      Carrier64_Faults_1 : Int := 238;
      Carrier64_Faults_2 : Int := 239;
      Carrier64_Faults_3 : Int := 240;
      Carrier65_Faults_0 : Int := 241;
      Carrier65_Faults_1 : Int := 242;
      Carrier65_Faults_2 : Int := 243;
      Carrier65_Faults_3 : Int := 244;
      Carrier66_Faults_0 : Int := 245;
      Carrier66_Faults_1 : Int := 246;
      Carrier66_Faults_2 : Int := 247;
      Carrier66_Faults_3 : Int := 248;
      Carrier67_Faults_0 : Int := 249;
      Carrier67_Faults_1 : Int := 250;
      Carrier67_Faults_2 : Int := 251;
      Carrier67_Faults_3 : Int := 252;
      Carrier68_Faults_0 : Int := 253;
      Carrier68_Faults_1 : Int := 254;
      Carrier68_Faults_2 : Int := 255;
      Carrier68_Faults_3 : Int := 256;
      Carrier69_Faults_0 : Int := 257;
      Carrier69_Faults_1 : Int := 258;
      Carrier69_Faults_2 : Int := 259;
      Carrier69_Faults_3 : Int := 260;
      Carrier70_Faults_0 : Int := 261;
      Carrier70_Faults_1 : Int := 262;
      Carrier70_Faults_2 : Int := 263;
      Carrier70_Faults_3 : Int := 264;
      Carrier71_Faults_0 : Int := 265;
      Carrier71_Faults_1 : Int := 266;
      Carrier71_Faults_2 : Int := 267;
      Carrier71_Faults_3 : Int := 268;
      Carrier72_Faults_0 : Int := 269;
      Carrier72_Faults_1 : Int := 270;
      Carrier72_Faults_2 : Int := 271;
      Carrier72_Faults_3 : Int := 272;
      Carrier73_Faults_0 : Int := 273;
      Carrier73_Faults_1 : Int := 274;
      Carrier73_Faults_2 : Int := 275;
      Carrier73_Faults_3 : Int := 276;
      Carrier74_Faults_0 : Int := 277;
      Carrier74_Faults_1 : Int := 278;
      Carrier74_Faults_2 : Int := 279;
      Carrier74_Faults_3 : Int := 280;
      Carrier75_Faults_0 : Int := 281;
      Carrier75_Faults_1 : Int := 282;
      Carrier75_Faults_2 : Int := 283;
      Carrier75_Faults_3 : Int := 284;
      Carrier76_Faults_0 : Int := 285;
      Carrier76_Faults_1 : Int := 286;
      Carrier76_Faults_2 : Int := 287;
      Carrier76_Faults_3 : Int := 288;
      Carrier77_Faults_0 : Int := 289;
      Carrier77_Faults_1 : Int := 290;
      Carrier77_Faults_2 : Int := 291;
      Carrier77_Faults_3 : Int := 292;
      Carrier78_Faults_0 : Int := 293;
      Carrier78_Faults_1 : Int := 294;
      Carrier78_Faults_2 : Int := 295;
      Carrier78_Faults_3 : Int := 296;
      Carrier79_Faults_0 : Int := 297;
      Carrier79_Faults_1 : Int := 298;
      Carrier79_Faults_2 : Int := 299;
      Carrier79_Faults_3 : Int := 300;
      Carrier80_Faults_0 : Int := 301;
      Carrier80_Faults_1 : Int := 302;
      Carrier80_Faults_2 : Int := 303;
      Carrier80_Faults_3 : Int := 304;
      Carrier81_Faults_0 : Int := 305;
      Carrier81_Faults_1 : Int := 306;
      Carrier81_Faults_2 : Int := 307;
      Carrier81_Faults_3 : Int := 308;
      Carrier82_Faults_0 : Int := 309;
      Carrier82_Faults_1 : Int := 310;
      Carrier82_Faults_2 : Int := 311;
      Carrier82_Faults_3 : Int := 312;
   END_VAR
BEGIN
END_DATA_BLOCK

DATA_BLOCK "DB401_HMI_Status"   // DB401
{ S7_Optimized_Access := 'TRUE' }
VERSION : 0.1
   VAR
      Drive : "UDT_Drive_HMI";
      IO : "UDT_Carrier_IO_HMI";
      Status : "UDT_Carrier_Status_HMI";
      ZoneStatus : "UDT_Zone_Status_HMI";
   END_VAR
BEGIN
END_DATA_BLOCK

DATA_BLOCK "DB402_SDC_CARRIER_DRIVE_DATA"   // DB402
{ S7_Optimized_Access := 'TRUE' }
VERSION : 0.1
   VAR
      Drive_Data : "UDT_Carrier_Drive_Data";
   END_VAR
BEGIN
END_DATA_BLOCK

DATA_BLOCK "DB403_SDC_CARRIER_IO"   // DB403
{ S7_Optimized_Access := 'TRUE' }
VERSION : 0.1
   VAR
      IO_Data : "UDT_Carrier_IO_Data";
   END_VAR
BEGIN
END_DATA_BLOCK

DATA_BLOCK "Data_block_DO_NOT_CHANGE"   // DB999
{ S7_Optimized_Access := 'TRUE' }
VERSION : 0.1
   VAR RETAIN
      Production_Spacing_Memory : Int := 1000;
      Carrier_Spacing_Memory : Int := 800;
   END_VAR
BEGIN
END_DATA_BLOCK

DATA_BLOCK "DB1000_AB_Interlocks"   // DB1000
{ S7_Optimized_Access := 'TRUE' }
VERSION : 0.1
   VAR
      Interlock : "UDT_AB_Interlocks";
   END_VAR
BEGIN
END_DATA_BLOCK

DATA_BLOCK "DB_SDC_GLOBAL"   // DB3700
{ S7_Optimized_Access := 'FALSE' }
AUTHOR : FFM
FAMILY : SDC
NAME : GLOBAL
VERSION : 1.0
   VAR
      EMS_ID_ACT : Int := 130;   // Aktuelle Anzahl der EMS-Treiber
      EMS_ID_MIN : Int := 1;   // Minimum EMS ID
      EMS_ID_MAX : Int := 184;   // Maximum EMS ID
      min_barcode_mm : DInt := 900;   // Lower limit, bar code value
      max_barcode_mm : DInt := 2076000;   // Upper limit, bar code value
      START_COURSE : DInt := 5800;   // Start Barcodevalue of Course
      END_COURSE : DInt := 312200;   // Ende Barcodewert vom Kurs
      SEK_MIN : Int := 1;   // Erste Abschnitt Nummer
      SEK_MAX : Int := 508;   // Aktuelle Anzahl der Bahnabschnitte
      TAKT_TIME : Int := 0;   // Reserve
      SEK_CYCLE_COUNTER : Int := 423;   // Section for increasing the track cycle counter
      MAN_V_1 : DInt := 6000;   // manual mode, set value: drive speed (mm/min)
      MAN_V_2 : DInt := 6000;   // manual mode, set value: drive speed (mm/min)
      min_Sequence_monitor_mm : DInt := 0;   // Lower limit of bar code value for sequence monitoring
      max_Sequence_monitor_mm : DInt := 0;   // Upper limit of bar code value for sequence monitoring
      MAX_PROFIL : Int := 10;   // maximal Profil Numbers
      CURR_EMS_ID_MAX : Int := 184;   // derzeit höchsten EMS-Nummer aktiv
      current_EMS_loop : Int := 0;   // Aktuelle Anzahl der EMS-Treiber auf Schleife
      EMS_ID_BUSY : Int := 0;   // EMS Driver wird aktiviert oder deaktiviert
      TAKT_TIME_LAST : Int := 0;   // Reserve
      Reserve_56 : Array[56..59] of Byte;
      SEK_REPAIR_1 : Int := 473;   // Section for repair, reset "send to repair 1" bit
      SEK_REPAIR_2 : Int := 0;   // Section for repair, reset "send to repair 2" bit
      SEK_DIAG_1 : Int := 0;   // Section diagnosticstation 1
      SEK_DIAG_2 : Int := 0;   // Section diagnosticstation 2
      SEK_DIAG_3 : Int := 0;   // Section diagnosticstation 2
      SEK_REP_1_START : Int := 470;
      SEK_REP_1_ENDE : Int := 472;
      SEK_REP_2_START : Int := 475;
      SEK_REP_2_ENDE : Int := 475;
      INFO_REP_1_DIAG_1 : Int := 0;   // Info for Function Rep 1 at Dignosticstation 1
      INFO_REP_2_DIAG_1 : Int := 0;   // Info for Function Rep 2 at Dignosticstation 1
      INFO_REP_1_DIAG_2 : Int := 0;   // Info for Function Rep 1 at Dignosticstation 2
      INFO_REP_2_DIAG_2 : Int := 0;   // Info for Function Rep 2 at Dignosticstation 2
      INFO_REP_1_DIAG_3 : Int := 0;   // Info for Function Rep 1 at Dignosticstation 2
      INFO_REP_2_DIAG_3 : Int := 0;   // Info for Function Rep 2 at Dignosticstation 2
      EMS_VCleaner_1 : Int := 0;   // EMS mit Vaccumreiniger No.1
      EMS_VCleaner_2 : Int := 0;   // EMS mit Vaccumreiniger No.2
      EMS_AKT_ZAEHLER_NR : Int := 131;   // EMS Aktualisierungsnummer
      EMS_AKT_ANZAHL : Int := 10;   // EMS Aktualisierunganzahl
      EMS_DIST_SEARCH : Int := 600;   // EMS Entfernungssuche zum vorderen EMS
      MIN_DIST_EMS : Array[0..15] of Int;   // minimum distance
      Reserve_132 : Array[132..149] of Byte;
      SYNCH : Array[0..15] of Struct   // Zur Abstandsregelung im Synchronbereich
         SET_DIST : Int;   // Set point value: distance (mm)
         SYNCH_DIST : Int;   // Start synchron distance value: distance (mm)
         HYST : Int;   // IO Hysterese
         K : Real;   // erreichen von Synchron Faktor
         MAX_FAKT : Real;   // Faktor für maximale Synchronisiergeschwindigkeit
         MIN_FAKT : Real;   // Faktor für minimale Synchronisiergeschwindigkeit
      END_STRUCT;
      Reserve_438 : Array[438..499] of Byte;   // spare
      LIMITS : Array[0..15] of Struct
         RAPID_SLOW : Int;   // Umstellung Begrenzung auf Abstand (mm), Einschränkung
         SLOW_SPEED_FAKT : Real;   // Faktor Geschwindigkeit für langsame Drehzahl
      END_STRUCT;
      Reserve_596 : Array[596..599] of Byte;   // spare
      "M" : Struct
         NEUSTART : Bool := FALSE;
         T_NEUSTART : Bool := FALSE;
         F_RESET : Bool := FALSE;
         "EMS_Read-Write" : Bool := FALSE;
         SDC_ER_Reset : Bool := FALSE;
      END_STRUCT;
   END_VAR
BEGIN
   MIN_DIST_EMS[0] := 6000;
   MIN_DIST_EMS[1] := 5970;
   MIN_DIST_EMS[2] := 6100;
   MIN_DIST_EMS[3] := 6000;
   MIN_DIST_EMS[4] := 6050;
   MIN_DIST_EMS[5] := 6100;
   MIN_DIST_EMS[6] := 6500;
   MIN_DIST_EMS[7] := 6500;
   MIN_DIST_EMS[8] := 6000;
   MIN_DIST_EMS[9] := 6250;
   MIN_DIST_EMS[10] := 6500;
   MIN_DIST_EMS[11] := 7000;
   MIN_DIST_EMS[12] := 7500;
   MIN_DIST_EMS[13] := 5950;
   MIN_DIST_EMS[14] := 5980;
   MIN_DIST_EMS[15] := 6500;
   SYNCH[0].SET_DIST := 6080;
   SYNCH[1].SET_DIST := 6030;
   SYNCH[2].SET_DIST := 6150;
   SYNCH[3].SET_DIST := 6080;
   SYNCH[4].SET_DIST := 6090;
   SYNCH[5].SET_DIST := 6400;
   SYNCH[6].SET_DIST := 6400;
   SYNCH[7].SET_DIST := 6400;
   SYNCH[8].SET_DIST := 6100;
   SYNCH[9].SET_DIST := 6300;
   SYNCH[10].SET_DIST := 6600;
   SYNCH[11].SET_DIST := 7100;
   SYNCH[12].SET_DIST := 7600;
   SYNCH[13].SET_DIST := 6510;
   SYNCH[14].SET_DIST := 6510;
   SYNCH[15].SET_DIST := 6510;
   SYNCH[0].SYNCH_DIST := 6400;
   SYNCH[1].SYNCH_DIST := 6450;
   SYNCH[2].SYNCH_DIST := 18000;
   SYNCH[3].SYNCH_DIST := 6200;
   SYNCH[4].SYNCH_DIST := 12000;
   SYNCH[5].SYNCH_DIST := 12000;
   SYNCH[6].SYNCH_DIST := 12000;
   SYNCH[7].SYNCH_DIST := 12000;
   SYNCH[8].SYNCH_DIST := 10000;
   SYNCH[9].SYNCH_DIST := 10000;
   SYNCH[10].SYNCH_DIST := 10000;
   SYNCH[11].SYNCH_DIST := 10000;
   SYNCH[12].SYNCH_DIST := 10000;
   SYNCH[13].SYNCH_DIST := 6800;
   SYNCH[14].SYNCH_DIST := 6800;
   SYNCH[15].SYNCH_DIST := 6800;
   SYNCH[0].HYST := 10;
   SYNCH[1].HYST := 4;
   SYNCH[2].HYST := 4;
   SYNCH[0].K := 1.0;
   SYNCH[1].K := 1.0;
   SYNCH[2].K := 1.0;
   SYNCH[3].K := 1.0;
   SYNCH[4].K := 1.3;
   SYNCH[5].K := 0.2;
   SYNCH[6].K := 0.2;
   SYNCH[7].K := 0.2;
   SYNCH[8].K := 1.0;
   SYNCH[9].K := 1.0;
   SYNCH[10].K := 1.0;
   SYNCH[11].K := 1.0;
   SYNCH[12].K := 1.0;
   SYNCH[13].K := 1.0;
   SYNCH[14].K := 1.0;
   SYNCH[15].K := 1.0;
   SYNCH[0].MAX_FAKT := 1.1;
   SYNCH[1].MAX_FAKT := 1.4;
   SYNCH[2].MAX_FAKT := 20.0;
   SYNCH[3].MAX_FAKT := 1.0;
   SYNCH[4].MAX_FAKT := 4.0;
   SYNCH[5].MAX_FAKT := 1.2;
   SYNCH[6].MAX_FAKT := 1.2;
   SYNCH[7].MAX_FAKT := 1.2;
   SYNCH[8].MAX_FAKT := 1.0;
   SYNCH[9].MAX_FAKT := 1.0;
   SYNCH[10].MAX_FAKT := 1.0;
   SYNCH[11].MAX_FAKT := 1.0;
   SYNCH[12].MAX_FAKT := 1.0;
   SYNCH[13].MAX_FAKT := 1.0;
   SYNCH[14].MAX_FAKT := 1.0;
   SYNCH[15].MAX_FAKT := 1.0;
   SYNCH[0].MIN_FAKT := 1.0;
   SYNCH[1].MIN_FAKT := 1.0;
   SYNCH[2].MIN_FAKT := 1.0;
   SYNCH[3].MIN_FAKT := 1.0;
   SYNCH[4].MIN_FAKT := 1.0;
   SYNCH[5].MIN_FAKT := 0.8;
   SYNCH[6].MIN_FAKT := 0.8;
   SYNCH[7].MIN_FAKT := 0.8;
   SYNCH[8].MIN_FAKT := 1.0;
   SYNCH[9].MIN_FAKT := 1.0;
   SYNCH[10].MIN_FAKT := 1.0;
   SYNCH[11].MIN_FAKT := 1.0;
   SYNCH[12].MIN_FAKT := 1.0;
   SYNCH[13].MIN_FAKT := 1.0;
   SYNCH[14].MIN_FAKT := 1.0;
   SYNCH[15].MIN_FAKT := 1.0;
   LIMITS[0].RAPID_SLOW := 7200;
   LIMITS[1].RAPID_SLOW := 7400;
   LIMITS[2].RAPID_SLOW := 7700;
   LIMITS[3].RAPID_SLOW := 8200;
   LIMITS[4].RAPID_SLOW := 8700;
   LIMITS[5].RAPID_SLOW := 6250;
   LIMITS[6].RAPID_SLOW := 7500;
   LIMITS[7].RAPID_SLOW := 7500;
   LIMITS[8].RAPID_SLOW := 6500;
   LIMITS[9].RAPID_SLOW := 6700;
   LIMITS[10].RAPID_SLOW := 7000;
   LIMITS[11].RAPID_SLOW := 7500;
   LIMITS[12].RAPID_SLOW := 8000;
   LIMITS[13].RAPID_SLOW := 6300;
   LIMITS[14].RAPID_SLOW := 6030;
   LIMITS[15].RAPID_SLOW := 7500;
   LIMITS[0].SLOW_SPEED_FAKT := 0.3;
   LIMITS[1].SLOW_SPEED_FAKT := 0.3;
   LIMITS[2].SLOW_SPEED_FAKT := 0.3;
   LIMITS[3].SLOW_SPEED_FAKT := 0.3;
   LIMITS[4].SLOW_SPEED_FAKT := 0.3;
   LIMITS[5].SLOW_SPEED_FAKT := 0.4;
   LIMITS[6].SLOW_SPEED_FAKT := 0.2;
   LIMITS[7].SLOW_SPEED_FAKT := 0.2;
   LIMITS[8].SLOW_SPEED_FAKT := 0.3;
   LIMITS[9].SLOW_SPEED_FAKT := 0.3;
   LIMITS[10].SLOW_SPEED_FAKT := 0.3;
   LIMITS[11].SLOW_SPEED_FAKT := 0.3;
   LIMITS[12].SLOW_SPEED_FAKT := 0.3;
   LIMITS[13].SLOW_SPEED_FAKT := 0.2;
   LIMITS[14].SLOW_SPEED_FAKT := 0.7;
   LIMITS[15].SLOW_SPEED_FAKT := 0.2;
   Reserve_132[132] := 16#00;
   Reserve_132[133] := 16#00;
   Reserve_132[134] := 16#00;
   Reserve_132[135] := 16#00;
   Reserve_132[136] := 16#00;
   Reserve_132[137] := 16#00;
   Reserve_132[138] := 16#00;
   Reserve_132[139] := 16#00;
   Reserve_132[140] := 16#00;
   Reserve_132[141] := 16#00;
   Reserve_132[142] := 16#00;
   Reserve_132[143] := 16#00;
   Reserve_132[144] := 16#00;
   Reserve_132[145] := 16#00;
   Reserve_132[146] := 16#00;
   Reserve_132[147] := 16#00;
   Reserve_132[148] := 16#00;
   Reserve_132[149] := 16#00;
   SYNCH[3].HYST := 4;
   SYNCH[4].HYST := 4;
   SYNCH[5].HYST := 0;
   SYNCH[6].HYST := 0;
   SYNCH[7].HYST := 0;
   SYNCH[8].HYST := 0;
   SYNCH[9].HYST := 0;
   SYNCH[10].HYST := 0;
   SYNCH[11].HYST := 0;
   SYNCH[12].HYST := 10;
   SYNCH[13].HYST := 4;
   SYNCH[14].HYST := 4;
   SYNCH[15].HYST := 4;
   Reserve_438[438] := 16#00;
   Reserve_438[439] := 16#00;
   Reserve_438[440] := 16#00;
   Reserve_438[441] := 16#00;
   Reserve_438[442] := 16#00;
   Reserve_438[443] := 16#00;
   Reserve_438[444] := 16#00;
   Reserve_438[445] := 16#00;
   Reserve_438[446] := 16#00;
   Reserve_438[447] := 16#00;
   Reserve_438[448] := 16#00;
   Reserve_438[449] := 16#00;
   Reserve_438[450] := 16#00;
   Reserve_438[451] := 16#00;
   Reserve_438[452] := 16#00;
   Reserve_438[453] := 16#00;
   Reserve_438[454] := 16#00;
   Reserve_438[455] := 16#00;
   Reserve_438[456] := 16#00;
   Reserve_438[457] := 16#00;
   Reserve_438[458] := 16#00;
   Reserve_438[459] := 16#00;
   Reserve_438[460] := 16#00;
   Reserve_438[461] := 16#00;
   Reserve_438[462] := 16#00;
   Reserve_438[463] := 16#00;
   Reserve_438[464] := 16#00;
   Reserve_438[465] := 16#00;
   Reserve_438[466] := 16#00;
   Reserve_438[467] := 16#00;
   Reserve_438[468] := 16#00;
   Reserve_438[469] := 16#00;
   Reserve_438[470] := 16#00;
   Reserve_438[471] := 16#00;
   Reserve_438[472] := 16#00;
   Reserve_438[473] := 16#00;
   Reserve_438[474] := 16#00;
   Reserve_438[475] := 16#00;
   // 32 more start values not shown
END_DATA_BLOCK

DATA_BLOCK "DB_SDC_EMS_FLAGS"   // DB3701
{ S7_Optimized_Access := 'FALSE' }
AUTHOR : FFM
FAMILY : SDC
NAME : GLOBAL
VERSION : 0.1
   VAR
      HEADER : Struct
         DB_NR : Int := 3701;
         MIN_NR_EMS : Int := 1;
         MAX_NR_EMS : Int := 200;
         START_EMS : Int := 20;
         LAENGE_EMS_FLAGS : Int := 2;
         ACT_COUNT : Int := 0;
         Res120 : Int := 0;
         Res140 : Int := 0;
         Res160 : Int := 0;
         Res180 : Int := 0;
      END_STRUCT;
      EMS : Array[1..200] of "UDT_SDC_EMS_FLAGS";
      LADDR_EMS : Array[1..200] of HW_ANY;
   END_VAR
BEGIN
   EMS[3].SIMULATION := FALSE;
   EMS[2].SIMULATION := FALSE;
   EMS[200].FAULTY := TRUE;
   EMS[199].FAULTY := TRUE;
   EMS[198].FAULTY := TRUE;
   EMS[197].FAULTY := TRUE;
   EMS[196].FAULTY := TRUE;
   EMS[195].FAULTY := TRUE;
   EMS[194].FAULTY := TRUE;
   EMS[193].FAULTY := TRUE;
   EMS[192].FAULTY := TRUE;
   EMS[191].FAULTY := TRUE;
   EMS[190].FAULTY := TRUE;
   EMS[189].FAULTY := TRUE;
   EMS[188].FAULTY := TRUE;
   EMS[187].FAULTY := TRUE;
   EMS[186].FAULTY := TRUE;
   EMS[185].FAULTY := TRUE;
   EMS[184].FAULTY := TRUE;
   EMS[183].FAULTY := TRUE;
   EMS[182].FAULTY := TRUE;
   EMS[181].FAULTY := TRUE;
   EMS[180].FAULTY := TRUE;
   EMS[179].FAULTY := TRUE;
   EMS[178].FAULTY := TRUE;
   EMS[177].FAULTY := TRUE;
   EMS[176].FAULTY := TRUE;
   EMS[175].FAULTY := TRUE;
   EMS[174].FAULTY := TRUE;
   EMS[173].FAULTY := TRUE;
   EMS[172].FAULTY := TRUE;
   EMS[171].FAULTY := TRUE;
   EMS[170].FAULTY := TRUE;
   EMS[169].FAULTY := TRUE;
   EMS[168].FAULTY := TRUE;
   EMS[167].FAULTY := TRUE;
   EMS[166].FAULTY := TRUE;
   EMS[165].FAULTY := TRUE;
   EMS[164].FAULTY := TRUE;
   EMS[163].FAULTY := TRUE;
   EMS[162].FAULTY := TRUE;
   EMS[161].FAULTY := TRUE;
   EMS[160].FAULTY := TRUE;
   EMS[159].FAULTY := TRUE;
   EMS[158].FAULTY := TRUE;
   EMS[157].FAULTY := TRUE;
   EMS[156].FAULTY := TRUE;
   EMS[155].FAULTY := TRUE;
   EMS[154].FAULTY := TRUE;
   EMS[153].FAULTY := TRUE;
   EMS[152].FAULTY := TRUE;
   EMS[151].FAULTY := TRUE;
   EMS[150].FAULTY := TRUE;
   EMS[149].FAULTY := TRUE;
   EMS[148].FAULTY := TRUE;
   EMS[147].FAULTY := TRUE;
   EMS[146].FAULTY := TRUE;
   EMS[145].FAULTY := TRUE;
   EMS[144].FAULTY := TRUE;
   EMS[143].FAULTY := TRUE;
   EMS[142].FAULTY := TRUE;
   EMS[141].FAULTY := TRUE;
   EMS[140].FAULTY := TRUE;
   EMS[139].FAULTY := TRUE;
   EMS[138].FAULTY := TRUE;
   EMS[137].FAULTY := TRUE;
   EMS[136].FAULTY := TRUE;
   EMS[135].FAULTY := TRUE;
   EMS[134].FAULTY := TRUE;
   EMS[133].FAULTY := TRUE;
   EMS[132].FAULTY := TRUE;
   EMS[131].FAULTY := TRUE;
   EMS[130].FAULTY := TRUE;
   EMS[129].FAULTY := TRUE;
   EMS[128].FAULTY := TRUE;
   EMS[127].FAULTY := TRUE;
   EMS[126].FAULTY := TRUE;
   EMS[125].FAULTY := TRUE;
   EMS[124].FAULTY := TRUE;
   EMS[123].FAULTY := TRUE;
   EMS[122].FAULTY := TRUE;
   EMS[121].FAULTY := TRUE;
   EMS[120].FAULTY := TRUE;
   EMS[119].FAULTY := TRUE;
   EMS[118].FAULTY := TRUE;
   EMS[117].FAULTY := TRUE;
   EMS[116].FAULTY := TRUE;
   EMS[115].FAULTY := TRUE;
   EMS[114].FAULTY := TRUE;
   EMS[113].FAULTY := TRUE;
   EMS[112].FAULTY := TRUE;
   EMS[111].FAULTY := TRUE;
   EMS[110].FAULTY := TRUE;
   EMS[109].FAULTY := TRUE;
   EMS[108].FAULTY := TRUE;
   EMS[107].FAULTY := TRUE;
   EMS[106].FAULTY := TRUE;
   EMS[105].FAULTY := TRUE;
   EMS[104].FAULTY := TRUE;
   EMS[103].FAULTY := TRUE;
   EMS[102].FAULTY := TRUE;
   EMS[101].FAULTY := TRUE;
   EMS[100].FAULTY := TRUE;
   EMS[99].FAULTY := TRUE;
   EMS[98].FAULTY := TRUE;
   EMS[97].FAULTY := TRUE;
   EMS[96].FAULTY := TRUE;
   EMS[95].FAULTY := TRUE;
   EMS[94].FAULTY := TRUE;
   EMS[93].FAULTY := TRUE;
   EMS[92].FAULTY := TRUE;
   EMS[91].FAULTY := TRUE;
   EMS[90].FAULTY := TRUE;
   EMS[89].FAULTY := TRUE;
   EMS[88].FAULTY := TRUE;
   EMS[87].FAULTY := TRUE;
   EMS[86].FAULTY := TRUE;
   EMS[85].FAULTY := TRUE;
   EMS[84].FAULTY := TRUE;
   EMS[83].FAULTY := TRUE;
   EMS[82].FAULTY := TRUE;
   EMS[81].FAULTY := TRUE;
   EMS[80].FAULTY := TRUE;
   EMS[79].FAULTY := TRUE;
   EMS[78].FAULTY := TRUE;
   EMS[77].FAULTY := TRUE;
   EMS[76].FAULTY := TRUE;
   EMS[75].FAULTY := TRUE;
   EMS[74].FAULTY := TRUE;
   EMS[73].FAULTY := TRUE;
   EMS[72].FAULTY := TRUE;
   EMS[71].FAULTY := TRUE;
   EMS[70].FAULTY := TRUE;
   EMS[69].FAULTY := TRUE;
   EMS[68].FAULTY := TRUE;
   EMS[67].FAULTY := TRUE;
   EMS[66].FAULTY := TRUE;
   EMS[65].FAULTY := TRUE;
   EMS[64].FAULTY := TRUE;
   EMS[63].FAULTY := TRUE;
   EMS[62].FAULTY := TRUE;
   EMS[61].FAULTY := TRUE;
   EMS[60].FAULTY := TRUE;
   EMS[59].FAULTY := TRUE;
   EMS[58].FAULTY := TRUE;
   EMS[57].FAULTY := TRUE;
   EMS[56].FAULTY := TRUE;
   EMS[55].FAULTY := TRUE;
   EMS[54].FAULTY := FALSE;
   EMS[53].FAULTY := TRUE;
   EMS[52].FAULTY := TRUE;
   EMS[51].FAULTY := TRUE;
   EMS[50].FAULTY := TRUE;
   EMS[49].FAULTY := TRUE;
   EMS[48].FAULTY := TRUE;
   EMS[47].FAULTY := TRUE;
   EMS[46].FAULTY := TRUE;
   EMS[45].FAULTY := TRUE;
   EMS[44].FAULTY := TRUE;
   EMS[43].FAULTY := TRUE;
   EMS[42].FAULTY := TRUE;
   EMS[41].FAULTY := TRUE;
   EMS[40].FAULTY := TRUE;
   EMS[39].FAULTY := TRUE;
   EMS[38].FAULTY := TRUE;
   EMS[37].FAULTY := TRUE;
   EMS[36].FAULTY := TRUE;
   EMS[35].FAULTY := TRUE;
   EMS[34].FAULTY := FALSE;
   EMS[33].FAULTY := TRUE;
   EMS[32].FAULTY := FALSE;
   EMS[31].FAULTY := TRUE;
   EMS[30].FAULTY := TRUE;
   EMS[29].FAULTY := FALSE;
   EMS[28].FAULTY := TRUE;
   EMS[27].FAULTY := TRUE;
   EMS[26].FAULTY := TRUE;
   EMS[25].FAULTY := TRUE;
   EMS[24].FAULTY := TRUE;
   EMS[23].FAULTY := TRUE;
   EMS[22].FAULTY := TRUE;
   EMS[21].FAULTY := TRUE;
   EMS[20].FAULTY := TRUE;
   EMS[19].FAULTY := TRUE;
   EMS[18].FAULTY := TRUE;
   EMS[17].FAULTY := TRUE;
   EMS[16].FAULTY := TRUE;
   EMS[15].FAULTY := TRUE;
   EMS[14].FAULTY := TRUE;
   EMS[13].FAULTY := TRUE;
   EMS[12].FAULTY := TRUE;
   EMS[11].FAULTY := TRUE;
   EMS[10].FAULTY := TRUE;
   EMS[9].FAULTY := TRUE;
   EMS[8].FAULTY := TRUE;
   EMS[7].FAULTY := TRUE;
   EMS[6].FAULTY := TRUE;
   EMS[5].FAULTY := TRUE;
   EMS[4].FAULTY := TRUE;
   EMS[3].FAULTY := TRUE;
   // 3200 more start values not shown
END_DATA_BLOCK

DATA_BLOCK "DB_SDC_TS_PARAMETER_1"   // DB3704
{ S7_Optimized_Access := 'FALSE' }
AUTHOR : FFM
FAMILY : SDC
NAME : SECT_DEF
VERSION : 1.0
   VAR
      HEADER : Struct
         DB_NR : Int := 3704;
         MIN_NR_SEK : Int := 1;
         MAX_NR_SEK : Int := 100;
         START_DAT : Int := 20;
         LAENGE_SEK_DATA : Int := 260;
         ANZ_PROFIL : Int := 10;
         OFFEST_PROFIL : Int := 40;
         LAENGE_PROFIL_DATA : Int := 22;
         Res160 : Int := 0;
         Res : Int := 0;
      END_STRUCT;
      TS : Array[1..100] of "UDT_SDC_TS_PARAMETER";
   END_VAR
BEGIN
   TS[100].ALLG.Drive_speed_2 := 15000;
   TS[100].ALLG.Drive_speed_1 := 15000;
   TS[100].ALLG.Stop_Position := 2674;
   TS[100].ALLG.POS.End_1 := 371999;
   TS[100].ALLG.POS.Start_1 := 365500;
   TS[96].ALLG.Drive_speed_2 := 10000;
   TS[96].ALLG.Drive_speed_1 := 15000;
   TS[96].ALLG.Stop_Position := 3000;
   TS[96].ALLG.POS.End_1 := 365499;
   TS[96].ALLG.POS.Start_1 := 357900;
   TS[95].ALLG.Drive_speed_2 := 10000;
   TS[95].ALLG.Drive_speed_1 := 15000;
   TS[95].ALLG.Stop_Position := 3000;
   TS[95].ALLG.POS.End_1 := 357899;
   TS[95].ALLG.POS.Start_1 := 351800;
   TS[94].ALLG.Drive_speed_2 := 10000;
   TS[94].ALLG.Drive_speed_1 := 15000;
   TS[94].ALLG.Stop_Position := 3000;
   TS[94].ALLG.POS.End_1 := 351799;
   TS[94].ALLG.POS.Start_1 := 345700;
   TS[93].ALLG.Drive_speed_2 := 10000;
   TS[93].ALLG.Drive_speed_1 := 15000;
   TS[93].ALLG.Stop_Position := 3000;
   TS[93].ALLG.POS.End_1 := 345699;
   TS[93].ALLG.POS.Start_1 := 339600;
   TS[92].ALLG.Drive_speed_2 := 10000;
   TS[92].ALLG.Drive_speed_1 := 15000;
   TS[92].ALLG.Stop_Position := 3000;
   TS[92].ALLG.POS.End_1 := 339599;
   TS[92].ALLG.POS.Start_1 := 333500;
   TS[91].ALLG.Drive_speed_2 := 10000;
   TS[91].ALLG.Drive_speed_1 := 15000;
   TS[91].ALLG.Stop_Position := 3000;
   TS[91].ALLG.POS.End_1 := 333499;
   TS[91].ALLG.POS.Start_1 := 327400;
   TS[90].ALLG.Drive_speed_2 := 10000;
   TS[90].ALLG.Drive_speed_1 := 15000;
   TS[90].ALLG.Stop_Position := 3000;
   TS[90].ALLG.POS.End_1 := 327399;
   TS[90].ALLG.POS.Start_1 := 321300;
   TS[89].ALLG.Drive_speed_2 := 10000;
   TS[89].ALLG.Drive_speed_1 := 15000;
   TS[89].ALLG.Stop_Position := 3000;
   TS[89].ALLG.POS.End_1 := 321299;
   TS[89].ALLG.POS.Start_1 := 315200;
   TS[88].ALLG.Drive_speed_2 := 10000;
   TS[88].ALLG.Drive_speed_1 := 15000;
   TS[88].ALLG.Stop_Position := 3000;
   TS[88].ALLG.POS.End_1 := 315199;
   TS[88].ALLG.POS.Start_1 := 309100;
   TS[87].ALLG.Drive_speed_2 := 10000;
   TS[87].ALLG.Drive_speed_1 := 15000;
   TS[87].ALLG.Stop_Position := 3000;
   TS[87].ALLG.POS.End_1 := 309099;
   TS[87].ALLG.POS.Start_1 := 303000;
   TS[86].ALLG.Drive_speed_2 := 10000;
   TS[86].ALLG.Drive_speed_1 := 15000;
   TS[86].ALLG.POS.End_1 := 302999;
   TS[86].ALLG.POS.Start_1 := 300000;
   TS[1].ALLG.SEK_NEXT_1 := 0;
   TS[1].ALLG.SEK_NEXT_2 := 0;
   TS[1].ALLG.Spare[4] := 16#00;
   TS[1].ALLG.Spare[5] := 16#00;
   TS[1].ALLG.POS.Start_1 := 1687400;
   TS[1].ALLG.POS.End_1 := 1693799;
   TS[1].ALLG.POS.Start_2 := 0;
   TS[1].ALLG.POS.End_2 := 0;
   TS[1].ALLG.POS.Actionpoint_1 := 0;
   TS[1].ALLG.POS.Actionpoint_2 := 0;
   TS[1].ALLG.FLAGS.DIST_VAL[0] := FALSE;
   TS[1].ALLG.FLAGS.DIST_VAL[1] := FALSE;
   TS[1].ALLG.FLAGS.DIST_VAL[2] := FALSE;
   TS[1].ALLG.FLAGS.DIST_VAL[3] := FALSE;
   TS[1].ALLG.FLAGS.DIST_VAL[4] := FALSE;
   TS[1].ALLG.FLAGS.DIST_VAL[5] := FALSE;
   TS[1].ALLG.FLAGS.DIST_VAL[6] := FALSE;
   TS[1].ALLG.FLAGS.DIST_VAL[7] := FALSE;
   TS[1].ALLG.FLAGS.DIST_VAL[8] := FALSE;
   TS[1].ALLG.FLAGS.DIST_VAL[9] := TRUE;
   TS[1].ALLG.FLAGS.DIST_VAL[10] := FALSE;
   TS[1].ALLG.FLAGS.DIST_VAL[11] := FALSE;
   TS[1].ALLG.FLAGS.DIST_VAL[12] := FALSE;
   TS[1].ALLG.FLAGS.DIST_VAL[13] := FALSE;
   TS[1].ALLG.FLAGS.DIST_VAL[14] := FALSE;
   TS[1].ALLG.FLAGS.DIST_VAL[15] := FALSE;
   TS[1].ALLG.FLAGS.one_profile := FALSE;
   TS[1].ALLG.FLAGS.BLIND := FALSE;
   TS[1].ALLG.FLAGS.NO_DIST_CONT := FALSE;
   TS[1].ALLG.FLAGS.SYNCH_AREA := FALSE;
   TS[1].ALLG.FLAGS.bit24 := FALSE;
   TS[1].ALLG.FLAGS.bit25 := FALSE;
   TS[1].ALLG.FLAGS.bit26 := FALSE;
   TS[1].ALLG.FLAGS.bit27 := FALSE;
   TS[1].ALLG.FLAGS.EN_HOIST := FALSE;
   TS[1].ALLG.FLAGS.D_RESET_AFTER := FALSE;
   TS[1].ALLG.FLAGS.D_PULK := FALSE;
   TS[1].ALLG.FLAGS.bit33 := FALSE;
   TS[1].ALLG.FLAGS.bit34 := FALSE;
   TS[1].ALLG.FLAGS.bit35 := FALSE;
   TS[1].ALLG.FLAGS.bit36 := FALSE;
   TS[1].ALLG.FLAGS.Deutronic_ON := FALSE;
   TS[1].ALLG.Stop_Position := 5800;
   TS[1].ALLG.Drive_speed_1 := 15000;
   TS[1].ALLG.Drive_speed_2 := 6000;
   TS[1].PROFIL[1].Hoist_Pos_start := 0;
   TS[1].PROFIL[1].Height := 3890;
   TS[1].PROFIL[1].Hoist_speed := 2000;
   TS[1].PROFIL[1].Hoist_offset_1 := 0;
   TS[1].PROFIL[1].Hoist_offset_2 := 0;
   TS[1].PROFIL[1].Hoist_offset_3 := 0;
   TS[1].PROFIL[1].Hoist_offset_4 := 0;
   TS[1].PROFIL[1].Hoist_Start_offset_1 := 0;
   TS[1].PROFIL[1].Hoist_Start_offset_2 := 0;
   TS[1].PROFIL[1].Hoist_Start_offset_3 := 0;
   TS[1].PROFIL[1].Hoist_Start_offset_4 := 0;
   TS[1].PROFIL[2].Hoist_Pos_start := 0;
   TS[1].PROFIL[2].Height := 3890;
   TS[1].PROFIL[2].Hoist_speed := 2000;
   TS[1].PROFIL[2].Hoist_offset_1 := 0;
   TS[1].PROFIL[2].Hoist_offset_2 := 0;
   TS[1].PROFIL[2].Hoist_offset_3 := 0;
   TS[1].PROFIL[2].Hoist_offset_4 := 0;
   TS[1].PROFIL[2].Hoist_Start_offset_1 := 0;
   TS[1].PROFIL[2].Hoist_Start_offset_2 := 0;
   TS[1].PROFIL[2].Hoist_Start_offset_3 := 0;
   TS[1].PROFIL[2].Hoist_Start_offset_4 := 0;
   TS[1].PROFIL[3].Hoist_Pos_start := 0;
   TS[1].PROFIL[3].Height := 3890;
   TS[1].PROFIL[3].Hoist_speed := 2000;
   TS[1].PROFIL[3].Hoist_offset_1 := 0;
   TS[1].PROFIL[3].Hoist_offset_2 := 0;
   TS[1].PROFIL[3].Hoist_offset_3 := 0;
   TS[1].PROFIL[3].Hoist_offset_4 := 0;
   TS[1].PROFIL[3].Hoist_Start_offset_1 := 0;
   TS[1].PROFIL[3].Hoist_Start_offset_2 := 0;
   TS[1].PROFIL[3].Hoist_Start_offset_3 := 0;
   TS[1].PROFIL[3].Hoist_Start_offset_4 := 0;
   TS[1].PROFIL[4].Hoist_Pos_start := 0;
   TS[1].PROFIL[4].Height := 3890;
   TS[1].PROFIL[4].Hoist_speed := 2000;
   TS[1].PROFIL[4].Hoist_offset_1 := 0;
   TS[1].PROFIL[4].Hoist_offset_2 := 0;
   TS[1].PROFIL[4].Hoist_offset_3 := 0;
   TS[1].PROFIL[4].Hoist_offset_4 := 0;
   TS[1].PROFIL[4].Hoist_Start_offset_1 := 0;
   TS[1].PROFIL[4].Hoist_Start_offset_2 := 0;
   TS[1].PROFIL[4].Hoist_Start_offset_3 := 0;
   TS[1].PROFIL[4].Hoist_Start_offset_4 := 0;
   TS[1].PROFIL[5].Hoist_Pos_start := 0;
   TS[1].PROFIL[5].Height := 3890;
   TS[1].PROFIL[5].Hoist_speed := 2000;
   TS[1].PROFIL[5].Hoist_offset_1 := 0;
   TS[1].PROFIL[5].Hoist_offset_2 := 0;
   TS[1].PROFIL[5].Hoist_offset_3 := 0;
   TS[1].PROFIL[5].Hoist_offset_4 := 0;
   TS[1].PROFIL[5].Hoist_Start_offset_1 := 0;
   TS[1].PROFIL[5].Hoist_Start_offset_2 := 0;
   TS[1].PROFIL[5].Hoist_Start_offset_3 := 0;
   TS[1].PROFIL[5].Hoist_Start_offset_4 := 0;
   TS[1].PROFIL[6].Hoist_Pos_start := 0;
   TS[1].PROFIL[6].Height := 3890;
   TS[1].PROFIL[6].Hoist_speed := 2000;
   TS[1].PROFIL[6].Hoist_offset_1 := 0;
   TS[1].PROFIL[6].Hoist_offset_2 := 0;
   TS[1].PROFIL[6].Hoist_offset_3 := 0;
   TS[1].PROFIL[6].Hoist_offset_4 := 0;
   TS[1].PROFIL[6].Hoist_Start_offset_1 := 0;
   TS[1].PROFIL[6].Hoist_Start_offset_2 := 0;
   TS[1].PROFIL[6].Hoist_Start_offset_3 := 0;
   TS[1].PROFIL[6].Hoist_Start_offset_4 := 0;
   TS[1].PROFIL[7].Hoist_Pos_start := 0;
   TS[1].PROFIL[7].Height := 3890;
   TS[1].PROFIL[7].Hoist_speed := 2000;
   TS[1].PROFIL[7].Hoist_offset_1 := 0;
   TS[1].PROFIL[7].Hoist_offset_2 := 0;
   TS[1].PROFIL[7].Hoist_offset_3 := 0;
   TS[1].PROFIL[7].Hoist_offset_4 := 0;
   TS[1].PROFIL[7].Hoist_Start_offset_1 := 0;
   TS[1].PROFIL[7].Hoist_Start_offset_2 := 0;
   TS[1].PROFIL[7].Hoist_Start_offset_3 := 0;
   TS[1].PROFIL[7].Hoist_Start_offset_4 := 0;
   TS[1].PROFIL[8].Hoist_Pos_start := 0;
   TS[1].PROFIL[8].Height := 3890;
   TS[1].PROFIL[8].Hoist_speed := 2000;
   TS[1].PROFIL[8].Hoist_offset_1 := 0;
   TS[1].PROFIL[8].Hoist_offset_2 := 0;
   TS[1].PROFIL[8].Hoist_offset_3 := 0;
   TS[1].PROFIL[8].Hoist_offset_4 := 0;
   TS[1].PROFIL[8].Hoist_Start_offset_1 := 0;
   TS[1].PROFIL[8].Hoist_Start_offset_2 := 0;
   TS[1].PROFIL[8].Hoist_Start_offset_3 := 0;
   TS[1].PROFIL[8].Hoist_Start_offset_4 := 0;
   TS[1].PROFIL[9].Hoist_Pos_start := 0;
   TS[1].PROFIL[9].Height := 3890;
   TS[1].PROFIL[9].Hoist_speed := 2000;
   TS[1].PROFIL[9].Hoist_offset_1 := 0;
   TS[1].PROFIL[9].Hoist_offset_2 := 0;
   TS[1].PROFIL[9].Hoist_offset_3 := 0;
   TS[1].PROFIL[9].Hoist_offset_4 := 0;
   TS[1].PROFIL[9].Hoist_Start_offset_1 := 0;
   // 15300 more start values not shown
END_DATA_BLOCK

DATA_BLOCK "DB_SDC_TS_PARAMETER_2"   // DB3705
{ S7_Optimized_Access := 'FALSE' }
AUTHOR : FFM
FAMILY : SDC
NAME : SECT_DEF
VERSION : 1.0
   VAR
      HEADER : Struct
         DB_NR : Int := 3705;
         MIN_NR_SEK : Int := 101;
         MAX_NR_SEK : Int := 200;
         START_DAT : Int := 20;
         LAENGE_SEK_DATA : Int := 260;
         ANZ_PROFIL : Int := 10;
         OFFEST_PROFIL : Int := 40;
         LAENGE_PROFIL_DATA : Int := 22;
         Res160 : Int := 0;
         Res : Int := 0;
      END_STRUCT;
      TS : Array[101..200] of "UDT_SDC_TS_PARAMETER";
   END_VAR
BEGIN
   TS[101].ALLG.POS.Start_1 := 372000;
   TS[101].ALLG.POS.End_1 := 378499;
   TS[101].ALLG.Stop_Position := 3000;
   TS[101].ALLG.Drive_speed_1 := 20000;
   TS[101].ALLG.Drive_speed_2 := 20000;
   TS[102].ALLG.POS.Start_1 := 378500;
   TS[102].ALLG.POS.End_1 := 384999;
   TS[102].ALLG.Stop_Position := 3000;
   TS[102].ALLG.Drive_speed_1 := 10000;
   TS[102].ALLG.Drive_speed_2 := 7000;
   TS[103].ALLG.POS.Start_1 := 385000;
   TS[103].ALLG.POS.End_1 := 391499;
   TS[103].ALLG.Stop_Position := 3000;
   TS[103].ALLG.Drive_speed_1 := 20000;
   TS[103].ALLG.Drive_speed_2 := 20000;
   TS[104].ALLG.POS.Start_1 := 391500;
   TS[104].ALLG.POS.End_1 := 397999;
   TS[104].ALLG.Stop_Position := 3000;
   TS[104].ALLG.Drive_speed_1 := 20000;
   TS[104].ALLG.Drive_speed_2 := 20000;
   TS[105].ALLG.POS.Start_1 := 398000;
   TS[105].ALLG.POS.End_1 := 404499;
   TS[105].ALLG.Stop_Position := 3000;
   TS[105].ALLG.Drive_speed_1 := 22000;
   TS[105].ALLG.Drive_speed_2 := 20000;
   TS[106].ALLG.POS.Start_1 := 404500;
   TS[106].ALLG.POS.End_1 := 410999;
   TS[106].ALLG.Stop_Position := 3000;
   TS[106].ALLG.Drive_speed_1 := 22000;
   TS[106].ALLG.Drive_speed_2 := 5000;
   TS[107].ALLG.POS.Start_1 := 411000;
   TS[107].ALLG.POS.End_1 := 417499;
   TS[107].ALLG.Stop_Position := 3000;
   TS[107].ALLG.Drive_speed_1 := 18000;
   TS[107].ALLG.Drive_speed_2 := 4000;
   TS[108].ALLG.POS.Start_1 := 417500;
   TS[108].ALLG.POS.End_1 := 423999;
   TS[108].ALLG.Stop_Position := 3000;
   TS[108].ALLG.Drive_speed_1 := 22000;
   TS[108].ALLG.Drive_speed_2 := 10000;
   TS[109].ALLG.POS.Start_1 := 424000;
   TS[109].ALLG.POS.End_1 := 430499;
   TS[109].ALLG.Stop_Position := 3000;
   TS[109].ALLG.Drive_speed_1 := 20000;
   TS[109].ALLG.Drive_speed_2 := 10000;
   TS[110].ALLG.POS.Start_1 := 430500;
   TS[110].ALLG.POS.End_1 := 436999;
   TS[110].ALLG.Stop_Position := 2674;
   TS[110].ALLG.Drive_speed_1 := 15000;
   TS[110].ALLG.Drive_speed_2 := 10000;
   TS[111].ALLG.POS.Start_1 := 437000;
   TS[111].ALLG.POS.End_1 := 443499;
   TS[111].ALLG.Stop_Position := 3000;
   TS[111].ALLG.Drive_speed_1 := 15000;
   TS[111].ALLG.Drive_speed_2 := 10000;
   TS[120].ALLG.POS.Start_1 := 443500;
   TS[120].ALLG.POS.End_1 := 450499;
   TS[120].ALLG.Stop_Position := 5200;
   TS[120].ALLG.Drive_speed_1 := 15000;
   TS[120].ALLG.Drive_speed_2 := 10000;
   TS[121].ALLG.POS.Start_1 := 450500;
   TS[121].ALLG.POS.End_1 := 457499;
   TS[121].ALLG.Stop_Position := 5500;
   TS[121].ALLG.Drive_speed_1 := 15000;
   TS[121].ALLG.Drive_speed_2 := 10000;
   TS[122].ALLG.POS.Start_1 := 457500;
   TS[122].ALLG.POS.End_1 := 463999;
   TS[122].ALLG.Stop_Position := 5000;
   TS[122].ALLG.Drive_speed_1 := 15000;
   TS[122].ALLG.Drive_speed_2 := 10000;
   TS[123].ALLG.POS.Start_1 := 464000;
   TS[123].ALLG.POS.End_1 := 470499;
   TS[123].ALLG.Stop_Position := 5100;
   TS[123].ALLG.Drive_speed_1 := 15000;
   TS[123].ALLG.Drive_speed_2 := 10000;
   TS[124].ALLG.POS.Start_1 := 470500;
   TS[124].ALLG.POS.End_1 := 476999;
   TS[124].ALLG.Stop_Position := 5000;
   TS[124].ALLG.Drive_speed_1 := 15000;
   TS[124].ALLG.Drive_speed_2 := 10000;
   TS[125].ALLG.POS.Start_1 := 477000;
   TS[125].ALLG.POS.End_1 := 483999;
   TS[125].ALLG.Stop_Position := 6400;
   TS[125].ALLG.Drive_speed_1 := 15000;
   TS[125].ALLG.Drive_speed_2 := 10000;
   TS[126].ALLG.POS.Start_1 := 484000;